   	SmartTags("DB_MouldEditor_HMI_uData_arShotSet{7}_Pressure{1}")=HiField(37,1)
   	SmartTags("DB_MouldEditor_HMI_uData_arShotSet{7}_Pressure{2}")=HiField(37,2)
   	SmartTags("DB_MouldEditor_HMI_uData_arShotSet{7}_Pressure{3}")=HiField(37,3)
   	SmartTags("DB_MouldEditor_HMI_uData_arShotSet{7}_Pressure{4}")=HiField(37,4)
   	SmartTags("DB_MouldEditor_HMI_uData_arShotSet{7}_Pressure{5}")=HiField(37,5)
   	SmartTags("DB_MouldEditor_HMI_uData_arShotSet{7}_Pressure{6}")=HiField(37,6)
   	
   	SmartTags("DB_MouldEditor_HMI_uData_arShotSet{8}_Pressure{1}")=HiField(42,1)
   	SmartTags("DB_MouldEditor_HMI_uData_arShotSet{8}_Pressure{2}")=HiField(42,2)
   	SmartTags("DB_MouldEditor_HMI_uData_arShotSet{8}_Pressure{3}")=HiField(42,3)
   	SmartTags("DB_MouldEditor_HMI_uData_arShotSet{8}_Pressure{4}")=HiField(42,4)
   	SmartTags("DB_MouldEditor_HMI_uData_arShotSet{8}_Pressure{5}")=HiField(42,5)
   	SmartTags("DB_MouldEditor_HMI_uData_arShotSet{8}_Pressure{6}")=HiField(42,6)
   	
   	'For PS = 2 To 37
   	'	Je = Int((5*PS)-1)
   	'	Flo = Int((5*PS)+1)
   	'	Pre = Int((5*PS)+2)
   	'SmartTags("DB_MouldEditor_HMI_uData_arShotSet{" & PS & "}_RefComponent") = HiField(Je,1)
   	'SmartTags("DB_MouldEditor_HMI_uData_arShotSet{" & PS & "}_MHNo") = HiField(Je,2)
   	'SmartTags("DB_MouldEditor_HMI_uData_arShotSet{" & PS & "}_FoamingTime") = HiField(Je,3)
   	'SmartTags("DB_MouldEditor_HMI_uData_sCalculatedValues_arTotalFlow{" & PS & "}") = HiField(Je,4)
   	'SmartTags("DB_MouldEditor_HMI_uData_arShotSet{" & PS & "}_PartWeight") = HiField(Je,5)
   	'SmartTags("DB_MouldEditor_HMI_uData_arShotSet{" & PS & "}_PartCounter") = HiField(Je,6)
   	'SmartTags("DB_MouldEditor_HMI_uData_arShotSet{" & PS & "}_PartShotDisable") = HiField(Je,7)
   	'SmartTags("DB_MouldEditor_HMI_uData_arShotSet{" & PS & "}_CPMoveAfterShot") = HiField(Je,8)
   	'SmartTags("DB_MouldEditor_HMI_uData_arShotSet{" & PS & "}_PurgeMHAfterShot") = HiField(Je,9)
   	'SmartTags("DB_MouldEditor_HMI_uData_arShotSet{"& PS &"}_Flow1")=HiField(Flo,1)
   	'SmartTags("DB_MouldEditor_HMI_uData_arShotSet{"& PS &"}_Flow{2}")=HiField(Flo,2)	
   	'SmartTags("DB_MouldEditor_HMI_uData_arShotSet{"& PS &"}_Flow{3}")=HiField(Flo,3)
   	'SmartTags("DB_MouldEditor_HMI_uData_arShotSet{"& PS &"}_Flow{4}")=HiField(Flo,4)
   	'SmartTags("DB_MouldEditor_HMI_uData_arShotSet{"& PS &"}_Flow{5}")=HiField(Flo,5)	
   	'SmartTags("DB_MouldEditor_HMI_uData_arShotSet{"& PS &"}_Flow{6}")=HiField(Flo,6)
   	'SmartTags("DB_MouldEditor_HMI_uData_arShotSet{"& PS &"}_Pressure{1}")=HiField(Pre,1)
   	'SmartTags("DB_MouldEditor_HMI_uData_arShotSet{"& PS &"}_Pressure{2}")=HiField(Pre,2)
   	'SmartTags("DB_MouldEditor_HMI_uData_arShotSet{"& PS &"}_Pressure{3}")=HiField(Pre,3)
   	'SmartTags("DB_MouldEditor_HMI_uData_arShotSet{"& PS &"}_Pressure{4}")=HiField(Pre,4)
   	'SmartTags("DB_MouldEditor_HMI_uData_arShotSet{"& PS &"}_Pressure{5}")=HiField(Pre,5)
   	'SmartTags("DB_MouldEditor_HMI_uData_arShotSet{"& PS &"}_Pressure{6}")=HiField(Pre,6)
   
   	'HmiRuntime.Screens("Tool Editor").ScreenItems("I/O field_4").ProcessValue=Je
   	'Next
   	
   	j = j + 1
   Loop
   
   'Close file
   f.Close
   Set f = Nothing
   
   SmartTags("ImportDataFrom_SD_stat")= 1
   
   bfde4b54-0db7-4817-8032-87127bf19bb9 "Readout of the data was successful!"
   
   'ReadData_1
   End If
   '// EOS //////////////////////////////////////////////////////////////////

VB script "FoamingAlarm"
   If SmartTags("DB919_ShotResultMach_ShotResult_Ma{0}_General_SendData") = True Then
   c82f6f27-c560-49f9-90e8-01e0a088b2a2 Foaming_Alarm,8
   c82f6f27-c560-49f9-90e8-01e0a088b2a2 Foaming_Alarm,9
   c82f6f27-c560-49f9-90e8-01e0a088b2a2 Foaming_Alarm,10
   
   
   'COMPONENT 1
   If SmartTags("DB919_ShotResultMach_ShotResult_Ma{0}_Component_Comp{1}_ComponentActive") = True Then
   	c82f6f27-c560-49f9-90e8-01e0a088b2a2 Foaming_Alarm,11
   End If
   
   'COMPONENT 2
   If SmartTags("DB919_ShotResultMach_ShotResult_Ma{0}_Component_Comp{2}_ComponentActive") = True Then
   	c82f6f27-c560-49f9-90e8-01e0a088b2a2 Foaming_Alarm,12
   End If
   
   'COMPONENT 3
   If SmartTags("DB919_ShotResultMach_ShotResult_Ma{0}_Component_Comp{3}_ComponentActive") = True Then
   	c82f6f27-c560-49f9-90e8-01e0a088b2a2 Foaming_Alarm,13
   End If
   
   'COMPONENT 4
   If SmartTags("DB919_ShotResultMach_ShotResult_Ma{0}_Component_Comp{4}_ComponentActive") = True Then
   	c82f6f27-c560-49f9-90e8-01e0a088b2a2 Foaming_Alarm,14
   End If
   'COMPONENT 5
   If SmartTags("DB919_ShotResultMach_ShotResult_Ma{0}_Component_Comp{5}_ComponentActive") = True Then
   	c82f6f27-c560-49f9-90e8-01e0a088b2a2 Foaming_Alarm,15
   End If
   'COMPONENT 6
   If SmartTags("DB919_ShotResultMach_ShotResult_Ma{0}_Component_Comp{6}_ComponentActive") = True Then
   	c82f6f27-c560-49f9-90e8-01e0a088b2a2 Foaming_Alarm,0
   End If
   'COMPONENT 7
   If SmartTags("DB919_ShotResultMach_ShotResult_Ma{0}_Component_Comp{7}_ComponentActive") = True Then
   	c82f6f27-c560-49f9-90e8-01e0a088b2a2 Foaming_Alarm,1
   End If
   'COMPONENT 8
   If SmartTags("DB919_ShotResultMach_ShotResult_Ma{0}_Component_Comp{8}_ComponentActive") = True Then
   	c82f6f27-c560-49f9-90e8-01e0a088b2a2 Foaming_Alarm,2
   End If
   End If

VB script "Save_TXT_File"
   Dim file, fso
    
    Set fso = CreateObject("Scripting.FileSystemObject")
    Set file = fso.CreateTextFile ("\Storage Card SD\SettingShiftPlan.txt", True)
    file.WriteLine(SmartTags("Shift1_Monday").Value)
    file.WriteLine(SmartTags("Shift2_Monday").Value)
   file.WriteLine(SmartTags("Shift3_Monday").Value)
   file.WriteLine(SmartTags("Shift4_Monday").Value)
   file.WriteLine(SmartTags("Shift1_Tuesday").Value)
    file.WriteLine(SmartTags("Shift2_Tuesday").Value)
    file.WriteLine(SmartTags("Shift3_Tuesday").Value)
    file.WriteLine(SmartTags("Shift4_Tuesday").Value)
    file.WriteLine(SmartTags("Shift1_Wenesday").Value)
     file.WriteLine(SmartTags("Shift2_Wenesday").Value) 
      file.WriteLine(SmartTags("Shift3_Wenesday").Value)
      file.WriteLine(SmartTags("Shift4_Wenesday").Value)
     file.WriteLine(SmartTags("Shift1_Thrusday").Value)
     file.WriteLine(SmartTags("Shift2_Thrusday").Value)
     file.WriteLine(SmartTags("Shift3_Thrusday").Value)
     file.WriteLine(SmartTags("Shift4_Thrusday").Value)
     file.WriteLine(SmartTags("Shift1_Friday").Value)
    file.WriteLine(SmartTags("Shift2_Friday").Value)
    file.WriteLine(SmartTags("Shift3_Friday").Value)
    file.WriteLine(SmartTags("Shift4_Friday").Value)
     file.WriteLine(SmartTags("Shift1_Saturday").Value)
       file.WriteLine(SmartTags("Shift2_Saturday").Value)
   file.WriteLine(SmartTags("Shift3_Saturday").Value)
    file.WriteLine(SmartTags("Shift4_Saturday").Value) 
     file.WriteLine(SmartTags("Shift1_Sunday").Value)
      file.WriteLine(SmartTags("Shift2_Sunday").Value)
      file.WriteLine(SmartTags("Shift3_Sunday").Value)
       file.WriteLine(SmartTags("Shift4_Sunday").Value)
      file.WriteLine(SmartTags("Check_Shift1_Monday").Value)
      file.WriteLine(SmartTags("Check_Shift2_Monday").Value)
      file.WriteLine(SmartTags("Check_Shift3_Monday").Value)
      file.WriteLine(SmartTags("Check_Shift4_Monday").Value)
     file.WriteLine(SmartTags("Check_Shift1_Tuesday").Value)
      file.WriteLine(SmartTags("Check_Shift2_Tuesday").Value)
      file.WriteLine(SmartTags("Check_Shift3_Tuesday").Value)
      file.WriteLine(SmartTags("Check_Shift4_Tuesday").Value)
    file.WriteLine(SmartTags("Check_Shift1_Wenesday").Value)
      file.WriteLine(SmartTags("Check_Shift2_Wenesday").Value)
      file.WriteLine(SmartTags("Check_Shift3_Wenesday").Value)
        file.WriteLine(SmartTags("Check_Shift4_Wenesday").Value) 
          file.WriteLine(SmartTags("Check_Shift1_Thrusday").Value)
     file.WriteLine(SmartTags("Check_Shift2_Thrusday").Value)
     file.WriteLine(SmartTags("Check_Shift3_Thrusday").Value)
      file.WriteLine(SmartTags("Check_Shift4_Thrusday").Value)
     file.WriteLine(SmartTags("Check_Shift1_Friday").Value)
     file.WriteLine(SmartTags("Check_Shift2_Friday").Value) 
      file.WriteLine(SmartTags("Check_Shift3_Friday").Value)
      file.WriteLine(SmartTags("Check_Shift4_Friday").Value)
      file.WriteLine(SmartTags("Check_Shift1_Saturday").Value)
      file.WriteLine(SmartTags("Check_Shift2_Saturday").Value)
      file.WriteLine(SmartTags("Check_Shift3_Saturday").Value)
    file.WriteLine(SmartTags("Check_Shift4_Saturday").Value)
     file.WriteLine(SmartTags("Check_Shift1_Sunday").Value)
     file.WriteLine(SmartTags("Check_Shift2_Sunday").Value)
     file.WriteLine(SmartTags("Check_Shift3_Sunday").Value)
      file.WriteLine(SmartTags("Check_Shift4_Sunday").Value)
     file.Close
    Set fso = Nothing
    Set file = Nothing  

VB script "MH_TestshotVisibility"
   If SmartTags("DB123_MH_IO_Signals_MH{0}_IN_MH_Auto_Mode")=True Or SmartTags("DB123_MH_IO_Signals_MH{0}_IN_MH_Manual_Mode")=True Then
   	HmiRuntime.Screens("0004_Mixinghead").ScreenItems("TesshotVisibility").Visible=False
   Else
   	HmiRuntime.Screens("0004_Mixinghead").ScreenItems("TesshotVisibility").Visible=true
   End If

VB script "RefreshAlarm"
   If  SmartTags("TP-Bereichszeiger_Picturenumber_Bildnummer")=24 And SmartTags("Alarm_Filter_Tag")= 10 Then
   	bec8f1e5-2ab1-45f6-ad91-1d37c469eb91 0024_ActualFaults,0
   	b21d3eaf-4e31-425c-ad1a-ba4e4002cacc Alarm_Filter_Tag,10
   ElseIf SmartTags("TP-Bereichszeiger_Picturenumber_Bildnummer")=24 And SmartTags("Alarm_Filter_Tag")= 11 Then
   	bec8f1e5-2ab1-45f6-ad91-1d37c469eb91 0024_ActualFaults,0
   	b21d3eaf-4e31-425c-ad1a-ba4e4002cacc Alarm_Filter_Tag,11
   
   ElseIf SmartTags("TP-Bereichszeiger_Picturenumber_Bildnummer")=24 And SmartTags("Alarm_Filter_Tag")= 12 Then
   	bec8f1e5-2ab1-45f6-ad91-1d37c469eb91 0024_ActualFaults,0
   	b21d3eaf-4e31-425c-ad1a-ba4e4002cacc Alarm_Filter_Tag,12
   
   ElseIf SmartTags("TP-Bereichszeiger_Picturenumber_Bildnummer")=24 And SmartTags("Alarm_Filter_Tag")= 13 Then
   	bec8f1e5-2ab1-45f6-ad91-1d37c469eb91 0024_ActualFaults,0
   	b21d3eaf-4e31-425c-ad1a-ba4e4002cacc Alarm_Filter_Tag,13
   			
   End If

VB script "Custom_Datalog"
   Dim fileName,folderName,fileLocation
   Dim fso,fctl,currentPosition,nextPosition,currentTime,dataValues
   
   fileName= Year(Now()) & "_"& Month(Now())
   folderName= "Storage Card USB\"
   fileLocation = folderName & fileName
   
   On Error Resume Next 
   
   		Set fso = CreateObject("FileCtl.FileSystem")
   		If (fso.Dir(folderName))= "" Then
   			fso.Mkdir folderName
   		End If
   		
   		If Err.Number<>0 Then
   			bfde4b54-0db7-4817-8032-87127bf19bb9 "Error # " & CStr(Err.Number) &" " &Err.Description&" " &Err.Source
   			Err.Clear
   		End If
   		
   		Set fctl = CreateObject("FileCtl.File")
   		fctl.Open fileLocation,8
   		
   		If Err.Number<>0 Then
   			bfde4b54-0db7-4817-8032-87127bf19bb9 "Error # " & CStr(Err.Number) &" " &Err.Description&" " &Err.Source
   			Err.Clear
   		End If
   		
   		currentPosition = fctl.Loc
   		nextPosition=fctl.Seek
   		
   		If currentPosition =1 And  nextPosition =1 Then
   			fctl.LinePrint "Time, Data Point 1, Data Point 2,Data Point 3, Data Point 4, Data Point 5"
   		End If
   		
   		currentTime = Hour(Time) & ":" & Minute(Time)
   		dataValues = currentTime & "01" &", "&"02"&","&"03"&","&"04"&","&"05"
   		fctl.LinePrint dataValues
   		fctl.Close
   		
   		bfde4b54-0db7-4817-8032-87127bf19bb9 CStr(fileLocation)

VB script "ReadDataFromUSB"
   '/////////////////////////////////////////////////////////////////////////
   ' en: Script for the readout of a text file      
   ' de: Skript zum Auslesen einer Textdatei
   ' Created: 29-05-2007
   ' Version: v0.1
   ' Author:  ZW										   only for Windows CE
   '/////////////////////////////////////////////////////////////////////////
   
   'Declaration of local tags - Deklaration von lokalen Variablen
   Dim f, path, MyZf, i, j, field, HiField(43,10), PS, Je, Flo, Pre
   
   'If bExtension = 0 Then
   	'path = "\flash\textfile.txt"
   '	path = "\Storage Card2\textfile.txt"
   'Else
   	'path = "\flash\textfile.csv"
   	path = SmartTags("ImportDataFrom_USB")'"\Storage Card USB"
   'End If
   
   'Error Routine - Fehlerroutine
   On Error Resume Next
   
   If SmartTags("ImportDataFrom_USB_stat")= 0 Then
   	'Create object - Objekt erstellen
   Set f = CreateObject("FileCtl.File")
   
   If Err.Number <> 0 Then
   	bfde4b54-0db7-4817-8032-87127bf19bb9 "Error #" & CStr(Err.Number) & " " & Err.Description
   	Err.Clear
   	Exit Sub
   End If
   
   'Open file - Datei öffnen
   f.open path, 1
   
   If Err.Number <> 0 Then
   	bfde4b54-0db7-4817-8032-87127bf19bb9 "Error #" & CStr(Err.Number) & " " & Err.Description
   	Err.Clear
   	Exit Sub
   End If
   
   'Loop
   Do While f.EOF = False
   	MyZf = f.LineInputString
   	field = Split(MyZf, ";")
   	
   	For i=0 To 43
   		field(i) = Replace(field(i), " ", "")
   		HiField(j,i) = field(i)
   	Next
   	
   	SmartTags("DB_MouldEditor_HMI_uData_uTools_tool_name") = HiField(1,1)
   	SmartTags("DB_MouldEditor_HMI_uData_uTools_PartShot_Amount") = HiField(2,1)
   	
   	SmartTags("DB_MouldEditor_HMI_uData_arShotSet{1}_RefComponent") = HiField(4,1)
   	SmartTags("DB_MouldEditor_HMI_uData_arShotSet{1}_MHNo") = HiField(4,2)
   	SmartTags("DB_MouldEditor_HMI_uData_arShotSet{1}_FoamingTime") = HiField(4,3)
   	SmartTags("DB_MouldEditor_HMI_uData_sCalculatedValues_arTotalFlow{1}") = HiField(4,4)
   	SmartTags("DB_MouldEditor_HMI_uData_arShotSet{1}_PartWeight") = HiField(4,5)
   	SmartTags("DB_MouldEditor_HMI_uData_arShotSet{1}_PartCounter") = HiField(4,6)
   	SmartTags("DB_MouldEditor_HMI_uData_arShotSet{1}_PartShotDisable") = HiField(4,7)
   	SmartTags("DB_MouldEditor_HMI_uData_arShotSet{1}_CPMoveAfterShot") = HiField(4,8)
   	SmartTags("DB_MouldEditor_HMI_uData_arShotSet{1}_PurgeMHAfterShot") = HiField(4,9)
   	
   	SmartTags("DB_MouldEditor_HMI_uData_arShotSet{2}_RefComponent") = HiField(9,1)
   	SmartTags("DB_MouldEditor_HMI_uData_arShotSet{2}_MHNo") = HiField(9,2)
   	SmartTags("DB_MouldEditor_HMI_uData_arShotSet{2}_FoamingTime") = HiField(9,3)
   	SmartTags("DB_MouldEditor_HMI_uData_sCalculatedValues_arTotalFlow{2}") = HiField(9,4)
   	SmartTags("DB_MouldEditor_HMI_uData_arShotSet{2}_PartWeight") = HiField(9,5)
   	SmartTags("DB_MouldEditor_HMI_uData_arShotSet{2}_PartCounter") = HiField(9,6)
   	SmartTags("DB_MouldEditor_HMI_uData_arShotSet{2}_PartShotDisable") = HiField(9,7)
   	SmartTags("DB_MouldEditor_HMI_uData_arShotSet{2}_CPMoveAfterShot") = HiField(9,8)
   	SmartTags("DB_MouldEditor_HMI_uData_arShotSet{2}_PurgeMHAfterShot") = HiField(9,9)
   	
   	SmartTags("DB_MouldEditor_HMI_uData_arShotSet{3}_RefComponent") = HiField(14,1)
   	SmartTags("DB_MouldEditor_HMI_uData_arShotSet{3}_MHNo") = HiField(14,2)
   	SmartTags("DB_MouldEditor_HMI_uData_arShotSet{3}_FoamingTime") = HiField(14,3)
   	SmartTags("DB_MouldEditor_HMI_uData_sCalculatedValues_arTotalFlow{3}") = HiField(14,4)
   	SmartTags("DB_MouldEditor_HMI_uData_arShotSet{3}_PartWeight") = HiField(14,5)
   	SmartTags("DB_MouldEditor_HMI_uData_arShotSet{3}_PartCounter") = HiField(14,6)
   	SmartTags("DB_MouldEditor_HMI_uData_arShotSet{3}_PartShotDisable") = HiField(14,7)
   	SmartTags("DB_MouldEditor_HMI_uData_arShotSet{3}_CPMoveAfterShot") = HiField(14,8)
   	SmartTags("DB_MouldEditor_HMI_uData_arShotSet{3}_PurgeMHAfterShot") = HiField(14,9)
   	
   	SmartTags("DB_MouldEditor_HMI_uData_arShotSet{4}_RefComponent") = HiField(19,1)
   	SmartTags("DB_MouldEditor_HMI_uData_arShotSet{4}_MHNo") = HiField(19,2)
   	SmartTags("DB_MouldEditor_HMI_uData_arShotSet{4}_FoamingTime") = HiField(19,3)
   	SmartTags("DB_MouldEditor_HMI_uData_sCalculatedValues_arTotalFlow{4}") = HiField(19,4)
   	SmartTags("DB_MouldEditor_HMI_uData_arShotSet{4}_PartWeight") = HiField(19,5)
   	SmartTags("DB_MouldEditor_HMI_uData_arShotSet{4}_PartCounter") = HiField(19,6)
   	SmartTags("DB_MouldEditor_HMI_uData_arShotSet{4}_PartShotDisable") = HiField(19,7)
   	SmartTags("DB_MouldEditor_HMI_uData_arShotSet{4}_CPMoveAfterShot") = HiField(19,8)
   	SmartTags("DB_MouldEditor_HMI_uData_arShotSet{4}_PurgeMHAfterShot") = HiField(19,9)
   	
   	SmartTags("DB_MouldEditor_HMI_uData_arShotSet{5}_RefComponent") = HiField(24,1)
   	SmartTags("DB_MouldEditor_HMI_uData_arShotSet{5}_MHNo") = HiField(24,2)
   	SmartTags("DB_MouldEditor_HMI_uData_arShotSet{5}_FoamingTime") = HiField(24,3)
   	SmartTags("DB_MouldEditor_HMI_uData_sCalculatedValues_arTotalFlow{5}") = HiField(24,4)
   	SmartTags("DB_MouldEditor_HMI_uData_arShotSet{5}_PartWeight") = HiField(24,5)
   	SmartTags("DB_MouldEditor_HMI_uData_arShotSet{5}_PartCounter") = HiField(24,6)
   	SmartTags("DB_MouldEditor_HMI_uData_arShotSet{5}_PartShotDisable") = HiField(24,7)
   	SmartTags("DB_MouldEditor_HMI_uData_arShotSet{5}_CPMoveAfterShot") = HiField(24,8)
   	SmartTags("DB_MouldEditor_HMI_uData_arShotSet{5}_PurgeMHAfterShot") = HiField(24,9)
   	
   	SmartTags("DB_MouldEditor_HMI_uData_arShotSet{6}_RefComponent") = HiField(29,1)
   	SmartTags("DB_MouldEditor_HMI_uData_arShotSet{6}_MHNo") = HiField(29,2)
   	SmartTags("DB_MouldEditor_HMI_uData_arShotSet{6}_FoamingTime") = HiField(29,3)
   	SmartTags("DB_MouldEditor_HMI_uData_sCalculatedValues_arTotalFlow{6}") = HiField(29,4)
   	SmartTags("DB_MouldEditor_HMI_uData_arShotSet{6}_PartWeight") = HiField(29,5)
   	SmartTags("DB_MouldEditor_HMI_uData_arShotSet{6}_PartCounter") = HiField(29,6)
   	SmartTags("DB_MouldEditor_HMI_uData_arShotSet{6}_PartShotDisable") = HiField(29,7)
   	SmartTags("DB_MouldEditor_HMI_uData_arShotSet{6}_CPMoveAfterShot") = HiField(29,8)
   	SmartTags("DB_MouldEditor_HMI_uData_arShotSet{6}_PurgeMHAfterShot") = HiField(29,9)
   	
   	SmartTags("DB_MouldEditor_HMI_uData_arShotSet{7}_RefComponent") = HiField(34,1)
   	SmartTags("DB_MouldEditor_HMI_uData_arShotSet{7}_MHNo") = HiField(34,2)
   	SmartTags("DB_MouldEditor_HMI_uData_arShotSet{7}_FoamingTime") = HiField(34,3)
   	SmartTags("DB_MouldEditor_HMI_uData_sCalculatedValues_arTotalFlow{7}") = HiField(34,4)
   	SmartTags("DB_MouldEditor_HMI_uData_arShotSet{7}_PartWeight") = HiField(34,5)
   	SmartTags("DB_MouldEditor_HMI_uData_arShotSet{7}_PartCounter") = HiField(34,6)
   	SmartTags("DB_MouldEditor_HMI_uData_arShotSet{7}_PartShotDisable") = HiField(34,7)
   	SmartTags("DB_MouldEditor_HMI_uData_arShotSet{7}_CPMoveAfterShot") = HiField(34,8)
   	SmartTags("DB_MouldEditor_HMI_uData_arShotSet{7}_PurgeMHAfterShot") = HiField(34,9)
   	
   	SmartTags("DB_MouldEditor_HMI_uData_arShotSet{8}_RefComponent") = HiField(39,1)
   	SmartTags("DB_MouldEditor_HMI_uData_arShotSet{8}_MHNo") = HiField(39,2)
   	SmartTags("DB_MouldEditor_HMI_uData_arShotSet{8}_FoamingTime") = HiField(39,3)
   	SmartTags("DB_MouldEditor_HMI_uData_sCalculatedValues_arTotalFlow{8}") = HiField(39,4)
   	SmartTags("DB_MouldEditor_HMI_uData_arShotSet{8}_PartWeight") = HiField(39,5)
   	SmartTags("DB_MouldEditor_HMI_uData_arShotSet{8}_PartCounter") = HiField(39,6)
   	SmartTags("DB_MouldEditor_HMI_uData_arShotSet{8}_PartShotDisable") = HiField(39,7)
   	SmartTags("DB_MouldEditor_HMI_uData_arShotSet{8}_CPMoveAfterShot") = HiField(39,8)
   	SmartTags("DB_MouldEditor_HMI_uData_arShotSet{8}_PurgeMHAfterShot") = HiField(39,9)
   	
   	'//FLOW
   	SmartTags("DB_MouldEditor_HMI_uData_arShotSet{1}_Flow{1}")=HiField(6,1)
   	SmartTags("DB_MouldEditor_HMI_uData_arShotSet{1}_Flow{2}")=HiField(6,2)	
   	SmartTags("DB_MouldEditor_HMI_uData_arShotSet{1}_Flow{3}")=HiField(6,3)
   	SmartTags("DB_MouldEditor_HMI_uData_arShotSet{1}_Flow{4}")=HiField(6,4)
   	SmartTags("DB_MouldEditor_HMI_uData_arShotSet{1}_Flow{5}")=HiField(6,5)	
   	SmartTags("DB_MouldEditor_HMI_uData_arShotSet{1}_Flow{6}")=HiField(6,6)
   	
   	SmartTags("DB_MouldEditor_HMI_uData_arShotSet{2}_Flow{1}")=HiField(11,1)
   	SmartTags("DB_MouldEditor_HMI_uData_arShotSet{2}_Flow{2}")=HiField(11,2)	
   	SmartTags("DB_MouldEditor_HMI_uData_arShotSet{2}_Flow{3}")=HiField(11,3)
   	SmartTags("DB_MouldEditor_HMI_uData_arShotSet{2}_Flow{4}")=HiField(11,4)
   	SmartTags("DB_MouldEditor_HMI_uData_arShotSet{2}_Flow{5}")=HiField(11,5)	
   	SmartTags("DB_MouldEditor_HMI_uData_arShotSet{2}_Flow{6}")=HiField(11,6)
   	
   	SmartTags("DB_MouldEditor_HMI_uData_arShotSet{3}_Flow{1}")=HiField(16,1)
   	SmartTags("DB_MouldEditor_HMI_uData_arShotSet{3}_Flow{2}")=HiField(16,2)	
   	SmartTags("DB_MouldEditor_HMI_uData_arShotSet{3}_Flow{3}")=HiField(16,3)
   	SmartTags("DB_MouldEditor_HMI_uData_arShotSet{3}_Flow{4}")=HiField(16,4)
   	SmartTags("DB_MouldEditor_HMI_uData_arShotSet{3}_Flow{5}")=HiField(16,5)	
   	SmartTags("DB_MouldEditor_HMI_uData_arShotSet{3}_Flow{6}")=HiField(16,6)
   	
   	SmartTags("DB_MouldEditor_HMI_uData_arShotSet{4}_Flow{1}")=HiField(21,1)
   	SmartTags("DB_MouldEditor_HMI_uData_arShotSet{4}_Flow{2}")=HiField(21,2)	
   	SmartTags("DB_MouldEditor_HMI_uData_arShotSet{4}_Flow{3}")=HiField(21,3)
   	SmartTags("DB_MouldEditor_HMI_uData_arShotSet{4}_Flow{4}")=HiField(21,4)
   	SmartTags("DB_MouldEditor_HMI_uData_arShotSet{4}_Flow{5}")=HiField(21,5)	
   	SmartTags("DB_MouldEditor_HMI_uData_arShotSet{4}_Flow{6}")=HiField(21,6)
   	
   	SmartTags("DB_MouldEditor_HMI_uData_arShotSet{5}_Flow{1}")=HiField(26,1)
   	SmartTags("DB_MouldEditor_HMI_uData_arShotSet{5}_Flow{2}")=HiField(26,2)	
   	SmartTags("DB_MouldEditor_HMI_uData_arShotSet{5}_Flow{3}")=HiField(26,3)
   	SmartTags("DB_MouldEditor_HMI_uData_arShotSet{5}_Flow{4}")=HiField(26,4)
   	SmartTags("DB_MouldEditor_HMI_uData_arShotSet{5}_Flow{5}")=HiField(26,5)	
   	SmartTags("DB_MouldEditor_HMI_uData_arShotSet{5}_Flow{6}")=HiField(26,6)
   	
   	SmartTags("DB_MouldEditor_HMI_uData_arShotSet{6}_Flow{1}")=HiField(31,1)
   	SmartTags("DB_MouldEditor_HMI_uData_arShotSet{6}_Flow{2}")=HiField(31,2)	
   	SmartTags("DB_MouldEditor_HMI_uData_arShotSet{6}_Flow{3}")=HiField(31,3)
   	SmartTags("DB_MouldEditor_HMI_uData_arShotSet{6}_Flow{4}")=HiField(31,4)
   	SmartTags("DB_MouldEditor_HMI_uData_arShotSet{6}_Flow{5}")=HiField(31,5)	
   	SmartTags("DB_MouldEditor_HMI_uData_arShotSet{6}_Flow{6}")=HiField(31,6)
   	
   	SmartTags("DB_MouldEditor_HMI_uData_arShotSet{7}_Flow{1}")=HiField(36,1)
   	SmartTags("DB_MouldEditor_HMI_uData_arShotSet{7}_Flow{2}")=HiField(36,2)	
   	SmartTags("DB_MouldEditor_HMI_uData_arShotSet{7}_Flow{3}")=HiField(36,3)
   	SmartTags("DB_MouldEditor_HMI_uData_arShotSet{7}_Flow{4}")=HiField(36,4)
   	SmartTags("DB_MouldEditor_HMI_uData_arShotSet{7}_Flow{5}")=HiField(36,5)	
   	SmartTags("DB_MouldEditor_HMI_uData_arShotSet{7}_Flow{6}")=HiField(36,6)
   	
   	SmartTags("DB_MouldEditor_HMI_uData_arShotSet{8}_Flow{1}")=HiField(41,1)
   	SmartTags("DB_MouldEditor_HMI_uData_arShotSet{8}_Flow{2}")=HiField(41,2)	
   	SmartTags("DB_MouldEditor_HMI_uData_arShotSet{8}_Flow{3}")=HiField(41,3)
   	SmartTags("DB_MouldEditor_HMI_uData_arShotSet{8}_Flow{4}")=HiField(41,4)
   	SmartTags("DB_MouldEditor_HMI_uData_arShotSet{8}_Flow{5}")=HiField(41,5)	
   	SmartTags("DB_MouldEditor_HMI_uData_arShotSet{8}_Flow{6}")=HiField(41,6)
   	
   	'//PRESSURE
   	SmartTags("DB_MouldEditor_HMI_uData_arShotSet{1}_Pressure{1}")=HiField(7,1)
   	SmartTags("DB_MouldEditor_HMI_uData_arShotSet{1}_Pressure{2}")=HiField(7,2)
   	SmartTags("DB_MouldEditor_HMI_uData_arShotSet{1}_Pressure{3}")=HiField(7,3)
   	SmartTags("DB_MouldEditor_HMI_uData_arShotSet{1}_Pressure{4}")=HiField(7,4)
   	SmartTags("DB_MouldEditor_HMI_uData_arShotSet{1}_Pressure{5}")=HiField(7,5)
   	SmartTags("DB_MouldEditor_HMI_uData_arShotSet{1}_Pressure{6}")=HiField(7,6)
   	
   	SmartTags("DB_MouldEditor_HMI_uData_arShotSet{2}_Pressure{1}")=HiField(12,1)
   	SmartTags("DB_MouldEditor_HMI_uData_arShotSet{2}_Pressure{2}")=HiField(12,2)
   	SmartTags("DB_MouldEditor_HMI_uData_arShotSet{2}_Pressure{3}")=HiField(12,3)
   	SmartTags("DB_MouldEditor_HMI_uData_arShotSet{2}_Pressure{4}")=HiField(12,4)
   	SmartTags("DB_MouldEditor_HMI_uData_arShotSet{2}_Pressure{5}")=HiField(12,5)
   	SmartTags("DB_MouldEditor_HMI_uData_arShotSet{2}_Pressure{6}")=HiField(12,6)
   	
   	SmartTags("DB_MouldEditor_HMI_uData_arShotSet{3}_Pressure{1}")=HiField(17,1)
   	SmartTags("DB_MouldEditor_HMI_uData_arShotSet{3}_Pressure{2}")=HiField(17,2)
   	SmartTags("DB_MouldEditor_HMI_uData_arShotSet{3}_Pressure{3}")=HiField(17,3)
   	SmartTags("DB_MouldEditor_HMI_uData_arShotSet{3}_Pressure{4}")=HiField(17,4)
   	SmartTags("DB_MouldEditor_HMI_uData_arShotSet{3}_Pressure{5}")=HiField(17,5)
   	SmartTags("DB_MouldEditor_HMI_uData_arShotSet{3}_Pressure{6}")=HiField(17,6)
   	
   	SmartTags("DB_MouldEditor_HMI_uData_arShotSet{4}_Pressure{1}")=HiField(22,1)
   	SmartTags("DB_MouldEditor_HMI_uData_arShotSet{4}_Pressure{2}")=HiField(22,2)
   	SmartTags("DB_MouldEditor_HMI_uData_arShotSet{4}_Pressure{3}")=HiField(22,3)
   	SmartTags("DB_MouldEditor_HMI_uData_arShotSet{4}_Pressure{4}")=HiField(22,4)
   	SmartTags("DB_MouldEditor_HMI_uData_arShotSet{4}_Pressure{5}")=HiField(22,5)
   	SmartTags("DB_MouldEditor_HMI_uData_arShotSet{4}_Pressure{6}")=HiField(22,6)
   	
   	SmartTags("DB_MouldEditor_HMI_uData_arShotSet{5}_Pressure{1}")=HiField(27,1)
   	SmartTags("DB_MouldEditor_HMI_uData_arShotSet{5}_Pressure{2}")=HiField(27,2)
   	SmartTags("DB_MouldEditor_HMI_uData_arShotSet{5}_Pressure{3}")=HiField(27,3)
   	SmartTags("DB_MouldEditor_HMI_uData_arShotSet{5}_Pressure{4}")=HiField(27,4)
   	SmartTags("DB_MouldEditor_HMI_uData_arShotSet{5}_Pressure{5}")=HiField(27,5)
   	SmartTags("DB_MouldEditor_HMI_uData_arShotSet{5}_Pressure{6}")=HiField(27,6)
   	
   	SmartTags("DB_MouldEditor_HMI_uData_arShotSet{6}_Pressure{1}")=HiField(32,1)
   	SmartTags("DB_MouldEditor_HMI_uData_arShotSet{6}_Pressure{2}")=HiField(32,2)
   	SmartTags("DB_MouldEditor_HMI_uData_arShotSet{6}_Pressure{3}")=HiField(32,3)
   	SmartTags("DB_MouldEditor_HMI_uData_arShotSet{6}_Pressure{4}")=HiField(32,4)
   	SmartTags("DB_MouldEditor_HMI_uData_arShotSet{6}_Pressure{5}")=HiField(32,5)
   	SmartTags("DB_MouldEditor_HMI_uData_arShotSet{6}_Pressure{6}")=HiField(32,6)
   	
   	SmartTags("DB_MouldEditor_HMI_uData_arShotSet{7}_Pressure{1}")=HiField(37,1)
   	SmartTags("DB_MouldEditor_HMI_uData_arShotSet{7}_Pressure{2}")=HiField(37,2)
   	SmartTags("DB_MouldEditor_HMI_uData_arShotSet{7}_Pressure{3}")=HiField(37,3)
   	SmartTags("DB_MouldEditor_HMI_uData_arShotSet{7}_Pressure{4}")=HiField(37,4)
   	SmartTags("DB_MouldEditor_HMI_uData_arShotSet{7}_Pressure{5}")=HiField(37,5)
   	SmartTags("DB_MouldEditor_HMI_uData_arShotSet{7}_Pressure{6}")=HiField(37,6)
   	
   	SmartTags("DB_MouldEditor_HMI_uData_arShotSet{8}_Pressure{1}")=HiField(42,1)
   	SmartTags("DB_MouldEditor_HMI_uData_arShotSet{8}_Pressure{2}")=HiField(42,2)
   	SmartTags("DB_MouldEditor_HMI_uData_arShotSet{8}_Pressure{3}")=HiField(42,3)
   	SmartTags("DB_MouldEditor_HMI_uData_arShotSet{8}_Pressure{4}")=HiField(42,4)
   	SmartTags("DB_MouldEditor_HMI_uData_arShotSet{8}_Pressure{5}")=HiField(42,5)
   	SmartTags("DB_MouldEditor_HMI_uData_arShotSet{8}_Pressure{6}")=HiField(42,6)
   	
   	'For PS = 2 To 37
   	'	Je = Int((5*PS)-1)
   	'	Flo = Int((5*PS)+1)
   	'	Pre = Int((5*PS)+2)
   	'SmartTags("DB_MouldEditor_HMI_uData_arShotSet{" & PS & "}_RefComponent") = HiField(Je,1)
   	'SmartTags("DB_MouldEditor_HMI_uData_arShotSet{" & PS & "}_MHNo") = HiField(Je,2)
   	'SmartTags("DB_MouldEditor_HMI_uData_arShotSet{" & PS & "}_FoamingTime") = HiField(Je,3)
   	'SmartTags("DB_MouldEditor_HMI_uData_sCalculatedValues_arTotalFlow{" & PS & "}") = HiField(Je,4)
   	'SmartTags("DB_MouldEditor_HMI_uData_arShotSet{" & PS & "}_PartWeight") = HiField(Je,5)
   	'SmartTags("DB_MouldEditor_HMI_uData_arShotSet{" & PS & "}_PartCounter") = HiField(Je,6)
   	'SmartTags("DB_MouldEditor_HMI_uData_arShotSet{" & PS & "}_PartShotDisable") = HiField(Je,7)
   	'SmartTags("DB_MouldEditor_HMI_uData_arShotSet{" & PS & "}_CPMoveAfterShot") = HiField(Je,8)
   	'SmartTags("DB_MouldEditor_HMI_uData_arShotSet{" & PS & "}_PurgeMHAfterShot") = HiField(Je,9)
   	'SmartTags("DB_MouldEditor_HMI_uData_arShotSet{"& PS &"}_Flow1")=HiField(Flo,1)
   	'SmartTags("DB_MouldEditor_HMI_uData_arShotSet{"& PS &"}_Flow{2}")=HiField(Flo,2)	
   	'SmartTags("DB_MouldEditor_HMI_uData_arShotSet{"& PS &"}_Flow{3}")=HiField(Flo,3)
   	'SmartTags("DB_MouldEditor_HMI_uData_arShotSet{"& PS &"}_Flow{4}")=HiField(Flo,4)
   	'SmartTags("DB_MouldEditor_HMI_uData_arShotSet{"& PS &"}_Flow{5}")=HiField(Flo,5)	
   	'SmartTags("DB_MouldEditor_HMI_uData_arShotSet{"& PS &"}_Flow{6}")=HiField(Flo,6)
   	'SmartTags("DB_MouldEditor_HMI_uData_arShotSet{"& PS &"}_Pressure{1}")=HiField(Pre,1)
   	'SmartTags("DB_MouldEditor_HMI_uData_arShotSet{"& PS &"}_Pressure{2}")=HiField(Pre,2)
   	'SmartTags("DB_MouldEditor_HMI_uData_arShotSet{"& PS &"}_Pressure{3}")=HiField(Pre,3)
   	'SmartTags("DB_MouldEditor_HMI_uData_arShotSet{"& PS &"}_Pressure{4}")=HiField(Pre,4)
   	'SmartTags("DB_MouldEditor_HMI_uData_arShotSet{"& PS &"}_Pressure{5}")=HiField(Pre,5)
   	'SmartTags("DB_MouldEditor_HMI_uData_arShotSet{"& PS &"}_Pressure{6}")=HiField(Pre,6)
   
   	'HmiRuntime.Screens("Tool Editor").ScreenItems("I/O field_4").ProcessValue=Je
   	'Next
   	
   	j = j + 1
   Loop
   
   'Close file
   f.Close
   Set f = Nothing
    SmartTags("ImportDataFrom_USB_stat")= 1
    
   bfde4b54-0db7-4817-8032-87127bf19bb9 "Readout of the data was successful!"
   
   'ReadData_1
   End If
   '// EOS //////////////////////////////////////////////////////////////////

VB script "Shift_Protocol"
   On Error Resume Next
   If SmartTags("CopyLogControl") <> 0 Then 'And Weekday = SmartTags("TP-Bereichszeiger_Date_Time_ActTime_WEEKDAY") And TimeValue(Now) = TimeValue(SmartTags("TP-Bereichszeiger_Date_Time_ActTime")) Then
   
   Select Case SmartTags("CopyLogControl")
   	Case 1
   		SmartTags("Shift_Protocol_21") = SmartTags("Shift_Protocol_20")
   		dd084c9b-3a0c-4857-9125-be72fcaad02d $3$hmiAlarmLog$, Schicht20, Schicht19, $3$hmiOverwrite$, $3$hmiYes$
   '		ShowSystemAlarm "Copy log success 21"
   	Case 2
   		SmartTags("Shift_Protocol_20") = SmartTags("Shift_Protocol_19")
   		dd084c9b-3a0c-4857-9125-be72fcaad02d $3$hmiAlarmLog$, Schicht19, Schicht18, $3$hmiOverwrite$, $3$hmiYes$
   '		ShowSystemAlarm "Copy log success 20"
   	Case 3
   		SmartTags("Shift_Protocol_19") = SmartTags("Shift_Protocol_18")
   		dd084c9b-3a0c-4857-9125-be72fcaad02d $3$hmiAlarmLog$, Schicht18, Schicht17, $3$hmiOverwrite$, $3$hmiYes$
   '		ShowSystemAlarm "Copy log success 19"
   	Case 4
   		SmartTags("Shift_Protocol_18") = SmartTags("Shift_Protocol_17")
   		dd084c9b-3a0c-4857-9125-be72fcaad02d $3$hmiAlarmLog$, Schicht17, Schicht16, $3$hmiOverwrite$, $3$hmiYes$
   '		ShowSystemAlarm "Copy log success 18"
   	Case 5
   		SmartTags("Shift_Protocol_17") = SmartTags("Shift_Protocol_16")
   		dd084c9b-3a0c-4857-9125-be72fcaad02d $3$hmiAlarmLog$, Schicht16, Schicht15, $3$hmiOverwrite$, $3$hmiYes$
   '		ShowSystemAlarm "Copy log success 17"
   	Case 6
   		SmartTags("Shift_Protocol_16") = SmartTags("Shift_Protocol_15")
   		dd084c9b-3a0c-4857-9125-be72fcaad02d $3$hmiAlarmLog$, Schicht15, Schicht14, $3$hmiOverwrite$, $3$hmiYes$
   '		ShowSystemAlarm "Copy log success 16"
   	Case 7
   		SmartTags("Shift_Protocol_15") = SmartTags("Shift_Protocol_14")
   		dd084c9b-3a0c-4857-9125-be72fcaad02d $3$hmiAlarmLog$, Schicht14, Schicht13, $3$hmiOverwrite$, $3$hmiYes$
   '		ShowSystemAlarm "Copy log success 15"
   	Case 8
   		SmartTags("Shift_Protocol_14") = SmartTags("Shift_Protocol_13")
   		dd084c9b-3a0c-4857-9125-be72fcaad02d $3$hmiAlarmLog$, Schicht13, Schicht12, $3$hmiOverwrite$, $3$hmiYes$
   '		ShowSystemAlarm "Copy log success 14"
   	Case 9
   		SmartTags("Shift_Protocol_13") = SmartTags("Shift_Protocol_12")
   		dd084c9b-3a0c-4857-9125-be72fcaad02d $3$hmiAlarmLog$, Schicht12, Schicht11, $3$hmiOverwrite$, $3$hmiYes$
   '		ShowSystemAlarm "Copy log success 13"
   	Case 10
   		SmartTags("Shift_Protocol_12") = SmartTags("Shift_Protocol_11")
   		dd084c9b-3a0c-4857-9125-be72fcaad02d $3$hmiAlarmLog$, Schicht11, Schicht10, $3$hmiOverwrite$, $3$hmiYes$
   '		ShowSystemAlarm "Copy log success 12"
   	Case 11
   		SmartTags("Shift_Protocol_11") = SmartTags("Shift_Protocol_10")
   		dd084c9b-3a0c-4857-9125-be72fcaad02d $3$hmiAlarmLog$, Schicht10, Schicht9, $3$hmiOverwrite$, $3$hmiYes$
   '		ShowSystemAlarm "Copy log success 11"
   	Case 12
   		SmartTags("Shift_Protocol_10") = SmartTags("Shift_Protocol_9")
   		dd084c9b-3a0c-4857-9125-be72fcaad02d $3$hmiAlarmLog$, Schicht9, Schicht8, $3$hmiOverwrite$, $3$hmiYes$
   '		ShowSystemAlarm "Copy log success 10"
   	Case 13
   		SmartTags("Shift_Protocol_9") = SmartTags("Shift_Protocol_8")
   		dd084c9b-3a0c-4857-9125-be72fcaad02d $3$hmiAlarmLog$, Schicht8, Schicht7, $3$hmiOverwrite$, $3$hmiYes$
   '		ShowSystemAlarm "Copy log success 9"
   	Case 14
   		SmartTags("Shift_Protocol_8") = SmartTags("Shift_Protocol_7")
   		dd084c9b-3a0c-4857-9125-be72fcaad02d $3$hmiAlarmLog$, Schicht7, Schicht6, $3$hmiOverwrite$, $3$hmiYes$
   '		ShowSystemAlarm "Copy log success 8"
   	Case 15
   		SmartTags("Shift_Protocol_7") = SmartTags("Shift_Protocol_6")
   		dd084c9b-3a0c-4857-9125-be72fcaad02d $3$hmiAlarmLog$, Schicht6, Schicht5, $3$hmiOverwrite$, $3$hmiYes$
   '		ShowSystemAlarm "Copy log success 7"
   	Case 16
   		SmartTags("Shift_Protocol_6") = SmartTags("Shift_Protocol_5")
   		dd084c9b-3a0c-4857-9125-be72fcaad02d $3$hmiAlarmLog$, Schicht5, Schicht4, $3$hmiOverwrite$, $3$hmiYes$
   '		ShowSystemAlarm "Copy log success 6"
   	Case 17
   		SmartTags("Shift_Protocol_5") = SmartTags("Shift_Protocol_4")
   		dd084c9b-3a0c-4857-9125-be72fcaad02d $3$hmiAlarmLog$, Schicht4, Schicht3, $3$hmiOverwrite$, $3$hmiYes$
   '		ShowSystemAlarm "Copy log success 5"
   	Case 18
   		SmartTags("Shift_Protocol_4") = SmartTags("Shift_Protocol_3")
   		dd084c9b-3a0c-4857-9125-be72fcaad02d $3$hmiAlarmLog$, Schicht3, Schicht2, $3$hmiOverwrite$, $3$hmiYes$
   '		ShowSystemAlarm "Copy log success 4"
   	Case 19
   		SmartTags("Shift_Protocol_3") = SmartTags("Shift_Protocol_2")
   		dd084c9b-3a0c-4857-9125-be72fcaad02d $3$hmiAlarmLog$, Schicht2, Schicht1, $3$hmiOverwrite$, $3$hmiYes$
   '		ShowSystemAlarm "Copy log success 3"
   	Case 20
   		SmartTags("Shift_Protocol_2") = SmartTags("Shift_Protocol_1")
   		dd084c9b-3a0c-4857-9125-be72fcaad02d $3$hmiAlarmLog$, Schicht1, Schicht0, $3$hmiOverwrite$, $3$hmiYes$
   '		ShowSystemAlarm "Copy log success 2"
   End Select
   End If
   If SmartTags("CopyLogControl") >= 21 Then
   	
   	SmartTags("Shift_Protocol_1") = SmartTags("Next shift")
   '	ShowSystemAlarm "Copy log success 1"
   	SettingShiftPlan
   	f38ba6b2-0c13-4a6f-acab-73f2fde9baea ShiftProtocol,1,$3$hmiOverwriteAlways$,$3$hmiOff$,Null	
   	SmartTags("CopyLogControl") = 0
   	
   End If
   	
   	

VB script "GetAlarmViewStat"
    HmiRuntime.Screens("0024_ActualFaults").ScreenItems("Pump Display Alarm").BackColor=vbBlue
    
    
    
    

VB script "CopyAlarmLogView"
   'SmartTags("CopyLogControl") = -1
   Select Case SmartTags("Archive Alarm Number")
   	Case 0
   		dd084c9b-3a0c-4857-9125-be72fcaad02d $3$hmiAlarmLog$,Archivanzeige,Schicht0,$3$hmiOverwrite$,$3$hmiNo$
   	Case 1
   		dd084c9b-3a0c-4857-9125-be72fcaad02d $3$hmiAlarmLog$,Archivanzeige,Schicht1,$3$hmiOverwrite$,$3$hmiNo$
   	Case 2
   		dd084c9b-3a0c-4857-9125-be72fcaad02d $3$hmiAlarmLog$,Archivanzeige,Schicht2,$3$hmiOverwrite$,$3$hmiNo$
   	Case 3
   		dd084c9b-3a0c-4857-9125-be72fcaad02d $3$hmiAlarmLog$,Archivanzeige,Schicht3,$3$hmiOverwrite$,$3$hmiNo$
   	Case 4
   		dd084c9b-3a0c-4857-9125-be72fcaad02d $3$hmiAlarmLog$,Archivanzeige,Schicht4,$3$hmiOverwrite$,$3$hmiNo$
   	Case 5
   		dd084c9b-3a0c-4857-9125-be72fcaad02d $3$hmiAlarmLog$,Archivanzeige,Schicht5,$3$hmiOverwrite$,$3$hmiNo$
   	Case 6
   		dd084c9b-3a0c-4857-9125-be72fcaad02d $3$hmiAlarmLog$,Archivanzeige,Schicht6,$3$hmiOverwrite$,$3$hmiNo$
   	Case 7
   		dd084c9b-3a0c-4857-9125-be72fcaad02d $3$hmiAlarmLog$,Archivanzeige,Schicht7,$3$hmiOverwrite$,$3$hmiNo$
   	Case 8
   		dd084c9b-3a0c-4857-9125-be72fcaad02d $3$hmiAlarmLog$,Archivanzeige,Schicht8,$3$hmiOverwrite$,$3$hmiNo$
   	Case 9
   		dd084c9b-3a0c-4857-9125-be72fcaad02d $3$hmiAlarmLog$,Archivanzeige,Schicht9,$3$hmiOverwrite$,$3$hmiNo$
   	Case 10
   		dd084c9b-3a0c-4857-9125-be72fcaad02d $3$hmiAlarmLog$,Archivanzeige,Schicht10,$3$hmiOverwrite$,$3$hmiNo$
   	Case 11
   		dd084c9b-3a0c-4857-9125-be72fcaad02d $3$hmiAlarmLog$,Archivanzeige,Schicht11,$3$hmiOverwrite$,$3$hmiNo$
   	Case 12
   		dd084c9b-3a0c-4857-9125-be72fcaad02d $3$hmiAlarmLog$,Archivanzeige,Schicht12,$3$hmiOverwrite$,$3$hmiNo$
   	Case 13
   		dd084c9b-3a0c-4857-9125-be72fcaad02d $3$hmiAlarmLog$,Archivanzeige,Schicht13,$3$hmiOverwrite$,$3$hmiNo$
   	Case 14
   		dd084c9b-3a0c-4857-9125-be72fcaad02d $3$hmiAlarmLog$,Archivanzeige,Schicht14,$3$hmiOverwrite$,$3$hmiNo$
   	Case 15
   		dd084c9b-3a0c-4857-9125-be72fcaad02d $3$hmiAlarmLog$,Archivanzeige,Schicht15,$3$hmiOverwrite$,$3$hmiNo$
   	Case 16
   		dd084c9b-3a0c-4857-9125-be72fcaad02d $3$hmiAlarmLog$,Archivanzeige,Schicht16,$3$hmiOverwrite$,$3$hmiNo$
   	Case 17
   		dd084c9b-3a0c-4857-9125-be72fcaad02d $3$hmiAlarmLog$,Archivanzeige,Schicht17,$3$hmiOverwrite$,$3$hmiNo$
   	Case 18
   		dd084c9b-3a0c-4857-9125-be72fcaad02d $3$hmiAlarmLog$,Archivanzeige,Schicht18,$3$hmiOverwrite$,$3$hmiNo$
   	Case 19
   		dd084c9b-3a0c-4857-9125-be72fcaad02d $3$hmiAlarmLog$,Archivanzeige,Schicht19,$3$hmiOverwrite$,$3$hmiNo$
   	Case 20
   		dd084c9b-3a0c-4857-9125-be72fcaad02d $3$hmiAlarmLog$,Archivanzeige,Schicht20,$3$hmiOverwrite$,$3$hmiNo$
   	Case 21
   		dd084c9b-3a0c-4857-9125-be72fcaad02d $3$hmiAlarmLog$,Archivanzeige,Schicht21,$3$hmiOverwrite$,$3$hmiNo$
   	
   End Select

VB script "EndShift"
   If Weekday(SmartTags("Next shift")) = SmartTags("TP-Bereichszeiger_Date_Time_ActTime_WEEKDAY") And Hour(SmartTags("Next shift")) = SmartTags("TP-Bereichszeiger_Date_Time_ActTime_HOUR") And Minute(SmartTags("Next shift")) = SmartTags("TP-Bereichszeiger_Date_Time_ActTime_MINUTE") And Second(SmartTags("Next shift")) = SmartTags("TP-Bereichszeiger_Date_Time_ActTime_SECOND") Then
   	b21d3eaf-4e31-425c-ad1a-ba4e4002cacc CopyLogControl,1
   	dd084c9b-3a0c-4857-9125-be72fcaad02d $3$hmiAlarmLog$,Schicht21,Schicht20,$3$hmiOverwrite$,$3$hmiYes$
   '	ShowSystemAlarm "Copy log 21 sukses"
   End If

VB script "Move_Act_Time"
   SmartTags("TP-Bereichszeiger_Date_Time_SetTime")=SmartTags("TP-Bereichszeiger_Date_Time_ActTime")

VB script "FirstScreen_NavigationUpdate"
   'SETTING PICTURE NAV 1 KIRI BERDASARKAN NOPAGE
   b21d3eaf-4e31-425c-ad1a-ba4e4002cacc Nav_1,SmartTags("DB14_TP_Shortcuts_TP_Shortcuts_PageNo_1")
   
   'SETTING PICTURE NAV 2 KIRI BERDASARKAN NOPAGE
   b21d3eaf-4e31-425c-ad1a-ba4e4002cacc Nav_2,SmartTags("DB14_TP_Shortcuts_TP_Shortcuts_PageNo_2")
   
   'SETTING PICTURE NAV 3 KIRI BERDASARKAN NOPAGE
   b21d3eaf-4e31-425c-ad1a-ba4e4002cacc Nav_3,SmartTags("DB14_TP_Shortcuts_TP_Shortcuts_PageNo_3")
   
   'SETTING PICTURE NAV 4 KIRI BERDASARKAN NOPAGE
   b21d3eaf-4e31-425c-ad1a-ba4e4002cacc Nav_4,SmartTags("DB14_TP_Shortcuts_TP_Shortcuts_PageNo_4")
   
   'SETTING PICTURE NAV 5 KIRI BERDASARKAN NOPAGE
   b21d3eaf-4e31-425c-ad1a-ba4e4002cacc Nav_5,SmartTags("DB14_TP_Shortcuts_TP_Shortcuts_PageNo_5")
   
   'SETTING PICTURE NAV 6 KIRI BERDASARKAN NOPAGE
   b21d3eaf-4e31-425c-ad1a-ba4e4002cacc Nav_6,SmartTags("DB14_TP_Shortcuts_TP_Shortcuts_PageNo_6")
   
   'SETTING PICTURE NAV 6 KIRI BERDASARKAN NOPAGE
   b21d3eaf-4e31-425c-ad1a-ba4e4002cacc Nav_7,SmartTags("DB14_TP_Shortcuts_TP_Shortcuts_PageNo_7")

VB script "Tes"
   Dim dtnow,sysnow,tnow,thnow,tmnow,tsnow,t1,t2,t3,th1,th2,th3,tm1,tm2,tm3,ts1,ts2,ts3
   dtnow=FormatDateTime(SmartTags("TP-Bereichszeiger_Date_Time_ActTime"),3)
   sysnow=FormatDateTime(Now(),3)
   
   
   thnow=Hour(dtnow)
   tmnow=Minute(dtnow)
   tsnow=Second(dtnow)
   
   tnow=FormatDateTime(SmartTags("TP-Bereichszeiger_Date_Time_ActTime"),3)
   t1=FormatDateTime(SmartTags("tes_Time_1"),3)
   t2=FormatDateTime(SmartTags("tes_Time_2"),3)
   t3=FormatDateTime(SmartTags("tes_Time_3"),3)
   
   th1=Hour(t1)
   tm1=Minute(t1)
   ts1=Second(t1)
   
   th2=Hour(t2)
   tm2=Minute(t2)
   ts2=Second(t2)
   
   th3=Hour(t3)
   tm3=Minute(t3)
   ts3=Second(t3)
   
   If sysnow<t1 Then
   	
   	SmartTags("tes_Time_3").Value=TimeSerial(CInt(th1),CInt(tm1),CInt(ts1))
   	
   ElseIf sysnow>t2 Then	
   	SmartTags("tes_Time_3").Value=TimeSerial(16,12,10)
   ElseIf sysnow<t2 And sysnow>t1 Then
   	SmartTags("tes_Time_3").Value=TimeSerial(CInt(th2),CInt(tm2),Cint(ts2))
   
   End If

VB script "SettingShiftPlan"
   Dim Shift, GT(8,4), NextS(4), Jam, Tanggal, WDay, N, Kosong, WeekD
   
   Jam = FormatDateTime(SmartTags("TP-Bereichszeiger_Date_Time_ActTime"),3)
   Tanggal = FormatDateTime(SmartTags("TP-Bereichszeiger_Date_Time_ActTime"),2)
   'Jam = FormatDateTime(Now,3)
   'Tanggal = FormatDateTime(Now,2)
   
   Kosong = 0
   
   If SmartTags("TP-Bereichszeiger_Date_Time_ActTime_WEEKDAY") > 1 Then
   	WeekD = (SmartTags("TP-Bereichszeiger_Date_Time_ActTime_WEEKDAY")-1)
   'If Weekday(Now) > 1 Then
   	'WeekD = (Weekday(Now)-1)
   Else
   	WeekD = 7
   End If
   
   For WDay = 1 To 7
   	For Shift = 1 To 4
   		If Not SmartTags("Shift_En_"& WDay & "_" & Shift) Then
   			GT(WDay,Shift) = "09/09/1999 09:09:00"
   		Else
   			Kosong = Kosong+1
   			If WDay = WeekD Then
   				If FormatDateTime(SmartTags("Shift_"& WDay & "_" & Shift),3) < Jam Then
   					GT(WDay,Shift) = "08/09/1999 " + FormatDateTime(SmartTags("Shift_"& WDay & "_" & Shift),3)
   				Else
   					GT(WDay,Shift) = SmartTags("Shift_"& WDay & "_" & Shift)
   				End If
   			End If
   			If WDay < WeekD Then
   				GT(WDay,Shift) = "07/09/1999 " + FormatDateTime(SmartTags("Shift_"& WDay & "_" & Shift),3)
   			End If
   			If WDay > WeekD Then
   				GT(WDay,Shift) = SmartTags("Shift_"& WDay & "_" & Shift)
   			End If
   		End If
   		'ShowSystemAlarm WDay & "_" & Shift & ": " & GT(WDay,Shift)
   	Next
   Next
   
   'On Error Resume Next
   For N = 7 To 1 Step -1
   If GT(N,1) < "02/02/1999 09:09:00" Or GT(N,2) < "02/02/1999 09:09:00" Or GT(N,3) < "02/02/1999 09:09:00" Or GT(N,4) < "02/02/1999 09:09:00" Then
   	WDay = N
   End If
   Next
   
   'ShowSystemAlarm "active day = " & WDay
   
   If WDay > 7 Then
   	For N = WeekD To 1 Step -1
   		If GT(N,1) <> "09/09/1999 09:09:00" Or GT(N,2) <> "09/09/1999 09:09:00" Or GT(N,3) <> "09/09/1999 09:09:00" Or GT(N,4) <> "09/09/1999 09:09:00" Then
   			WDay = N
   '			ShowSystemAlarm "active day = " & WDay
   		End If
   	Next
   End If
   
   'ShowSystemAlarm "active day = " & WDay
   
   If WDay >= WeekD Then
   	Tanggal = DateAdd("d",(WDay+1-(WeekD+1)),Tanggal)
   Else
   	Tanggal = DateAdd("d",(WDay+8-(WeekD+1)),Tanggal)
   End If
   
   'ShowSystemAlarm Tanggal
   	
   If GT(WDay,1) < GT(WDay,2) Then
   	NextS(1) = GT(WDay,1)
   Else
   	NextS(1) = GT(WDay,2)
   End If
   
   If GT(WDay,3) < GT(WDay,4) Then
   	NextS(2) = GT(WDay,3)
   Else
   	NextS(2) = GT(WDay,4)
   End If
   
   If NextS(1) < NextS(2) Then
   	SmartTags("Next shift") = (CDate(Tanggal) + TimeValue(FormatDateTime(NextS(1),3)))
   Else
   	SmartTags("Next shift") = (CDate(Tanggal) + TimeValue(FormatDateTime(NextS(2),3)))
   End If
   
   If WDay = WeekD And FormatDateTime(SmartTags("Next shift"),3) < Jam Then
   	SmartTags("Next shift") = DateAdd("d",7,SmartTags("Next shift"))
   End If
   
   If Kosong = 0 Then	
   	SmartTags("Next shift") = CDate("09/09/1999 09:09:00")
   End If
   
   'ShowSystemAlarm CStr(DateDiff("d",SmartTags("TP-Bereichszeiger_Date_Time_ActTime"),SmartTags("Next shift")))
   'ShowSystemAlarm CStr(SmartTags("Next shift"))
   'ShowSystemAlarm Jam

VB script "Shifttime_write"
   Dim fs, f, FName
   
   On Error Resume Next
    ' FileSystemObject erstellen
    ' Create FileSystemObject
   Set fs = CreateObject("FileCtl.FileSystem") 
   
   ' FileObject erstellen
   ' Create FileObject
    Set f = CreateObject("FileCtl.File")
    
   'FName = "Storage Card SD\Logs\Shifttime.txt" 
   FName = "Storage Card SD\Shifttime.txt" 
   
   
    f.open FName, 2								
   
    f.lineprint("Shift_1_1")
    f.lineprint("Shift_1_2")
    f.lineprint("Shift_1_3")
    f.lineprint("Shift_1_4")
    f.lineprint("Shift_2_1")
    f.lineprint("Shift_2_2")
    f.lineprint("Shift_2_3")
    f.lineprint("Shift_2_4")
    f.lineprint("Shift_3_1")
    f.lineprint("Shift_3_2")
    f.lineprint("Shift_3_3")
    f.lineprint("Shift_3_4") 
    f.lineprint("Shift_4_1")
    f.lineprint("Shift_4_2")
    f.lineprint("Shift_4_3")
    f.lineprint("Shift_4_4")
    f.lineprint("Shift_5_1")
    f.lineprint("Shift_5_2")
    f.lineprint("Shift_5_3")
    f.lineprint("Shift_5_4")
    f.lineprint("Shift_6_1")
    f.lineprint("Shift_6_2")
    f.lineprint("Shift_6_3")
    f.lineprint("Shift_6_4")
    f.lineprint("Shift_7_1")
    f.lineprint("Shift_7_2")
    f.lineprint("Shift_7_3")
    f.lineprint("Shift_7_4")
    f.lineprint("Shift_En_1_1")
    f.lineprint("Shift_En_1_2")
    f.lineprint("Shift_En_1_3")
    f.lineprint("Shift_En_1_4")
    f.lineprint("Shift_En_2_1")
    f.lineprint("Shift_En_2_2")
    f.lineprint("Shift_En_2_3")
    f.lineprint("Shift_En_2_4")
    f.lineprint("Shift_En_3_1")
    f.lineprint("Shift_En_3_2")
    f.lineprint("Shift_En_3_3")
    f.lineprint("Shift_En_3_4")
    f.lineprint("Shift_En_4_1")
    f.lineprint("Shift_En_4_2")
    f.lineprint("Shift_En_4_3")
    f.lineprint("Shift_En_4_4")
    f.lineprint("Shift_En_5_1")
    f.lineprint("Shift_En_5_2")
    f.lineprint("Shift_En_5_3")
    f.lineprint("Shift_En_5_4")
    f.lineprint("Shift_En_6_1")
    f.lineprint("Shift_En_6_2")
    f.lineprint("Shift_En_6_3")
    f.lineprint("Shift_En_6_4")
    f.lineprint("Shift_En_7_1")
    f.lineprint("Shift_En_7_2")
    f.lineprint("Shift_En_7_3")
    f.lineprint("Shift_En_7_4")
   ' Datei wieder schließen
   ' Close file
    f.Close
   Set f  = Nothing
   Set fs = Nothing
   'Error checking
   If Err.Number <>0 Then
   bfde4b54-0db7-4817-8032-87127bf19bb9 "Error#" & CStr(Err.Number) & " " & Err.Description
   Err.Clear
   ' Exit Sub'
   End If

VB script "Show_Not_Valid"
   If SmartTags("DB_MouldEditor_HMI_uData_sStatusBits_xFaultValuesnotvalid") = True Then
   	efd93a16-2665-4b85-bcb9-25eddcb7b6f4 Fault, 446, 387, $3$hmiOn$, $3$hmiAnimationOff$, $3$hmiMedium$
   Else
   	efd93a16-2665-4b85-bcb9-25eddcb7b6f4 Fault, 446, 387, $3$hmiOff$, $3$hmiAnimationOff$, $3$hmiMedium$
   End If

VB script "Read_USB_device"
   Dim fso,drive,result
   Set fso = CreateObject("Scripting.FileSystemObject")
   
   On Error Resume Next
   Set drive = fso.GetDrive(fso.GetDriveName(fso.GetAbsolutePathName(path)))
   
   If Err.Number = 0 Then
   	result = 0
   	bfde4b54-0db7-4817-8032-87127bf19bb9 "USB ADA !!!"
   	
   Else
   	result = Err.Number
   End If
   Read_USB_device = result

scheduled task "User_Change"
   on Action: function_e1ab61de("NavUserChange")
*)